HMI tags "Default tag table"
   "Tag_ScreenNumber" : UInt AT %DB1.DBW0
   "Part At Entry (NC)" : Bool AT %DB1.DBX0.0
   "InputsDB_Sensors_Part Entry" : Bool = PLC InputsDB.Sensors."Part Entry" AT %DB1.DBX0.0, 100 ms
   "Modes_Modes_RunMode" : Bool = PLC Modes.Modes.RunMode, 100 ms
   "HmiDb_ActivateUnloadHmi" : Bool = PLC HmiDb.HmiModes.ActivateUnloadHmi, 100 ms
   "Modes_Modes_StopMode" : Bool = PLC Modes.Modes.StoppestMode, 100 ms
   "Modes_Modes_ResetMode" : Bool = PLC Modes.Modes.ResetMode, 100 ms
   "HmiDb_HmiRunMode" : Bool = PLC HmiDb.HmiModes.HmiRunMode, 100 ms
   "HmiDb_HmiStopmode" : Bool = PLC HmiDb.HmiModes.HmiStopmode, 100 ms
   "HmiDb_HmiResetMode" : Bool = PLC HmiDb.HmiModes.HmiResetMode, 100 ms
   "InputsDB_Sensors_Part Load" : Bool = PLC InputsDB.Sensors."Part Load", 100 ms
   "InputsDB_Sensors_Part Unload" : Bool = PLC InputsDB.Sensors."Part Unload", 100 ms
   "InputsDB_Sensors_Part Exit" : Bool = PLC InputsDB.Sensors."Part Exit", 100 ms
   "InputsDB_Sensors_Crane Default" : Bool = PLC InputsDB.Sensors."Crane Default", 100 ms
   "InputsDB_Sensors_Crane Entry" : Bool = PLC InputsDB.Sensors."Crane Entry", 100 ms
   "InputsDB_Sensors_Color Sensor" : Int = PLC InputsDB.Sensors."Color Sensor", 100 ms
   "Modes_SafetyStops_ProductionStop" : Bool = PLC Modes.StopMethods.ProductionStop, 100 ms
   "Modes_SafetyStops_SafetyStop" : Bool = PLC Modes.StopMethods.SafetyStop, 100 ms
   "alarmStuck" : Int = PLC alarmStuck AT %QW34, 100 ms
   "alarmreceivedstuck" : UInt, internal
   "alarmLoaderFull" : Int = PLC alarmLoaderFull AT %QW36, 100 ms
   "alarmUnloaderEmpty" : Int = PLC alarmUnloaderEmpty AT %QW38, 100 ms
   "Modes_JogMode" : Bool = PLC Modes.Modes.JogMode, 100 ms
   "HmiDb_HmiRunEntryConv" : Bool = PLC HmiDb.ActivateAcutator.HmiRunEntryConv, 100 ms
   "HmiDb_HmiRunExitConv" : Bool = PLC HmiDb.ActivateAcutator.HmiRunExitConv, 100 ms
   "EntryConv" : Int = PLC InputsDB.ConvertedConveyors.EntryConvSensorVal, 100 ms
   "LoadingConv" : Int = PLC InputsDB.ConvertedConveyors.LoadingConvSensorVal, 100 ms
   "UnloadingConv" : Int = PLC InputsDB.ConvertedConveyors.UnloadingSensorVal, 100 ms
   "ExitConv" : Int = PLC InputsDB.ConvertedConveyors.ExitConvSensorVal, 100 ms
   "ohioselecter" : Int AT %DB1.DBW0
   "unloadingms" : Real = PLC InputsDB.ConvertedConveyors.UnloadingScaleX, 100 ms
   "loadingms" : Real = PLC InputsDB.ConvertedConveyors.LoadingConvScalex, 100 ms
   "exitms" : Real = PLC InputsDB.ConvertedConveyors.ExitConvScaleX, 100 ms
   "entryms" : Real = PLC InputsDB.ConvertedConveyors.EntryConvScalex, 100 ms
   "OutputsDB_CraneOutput_XScalex" : Int = PLC OutputsDB.CraneOutput.Xmm, 100 ms
   "OutputsDB_CraneOutput_YScalex" : Int = PLC OutputsDB.CraneOutput.Ymm, 100 ms
   "HmiDb_HmiExtendExit" : Bool = PLC HmiDb.ActivateAcutator.HmiExtendExit, 100 ms
   "HmiDb_HmiExtendEntry" : Bool = PLC HmiDb.ActivateAcutator.HmiExtendEntry, 100 ms
   "InputsDB_Sensors_Crane Exit" : Bool = PLC InputsDB.Sensors."Crane Exit", 100 ms
   "InputsDB_ConveyorCalibrationBarSlider" : Int = PLC InputsDB.ConveyorCalibrationBarSlider, 100 ms
   "InputsDB_ConveyorCalibrationPicker" : Int = PLC InputsDB.ConveyorCalibrationPicker, 100 ms
   "InputsDB_ConveyorSaveCalVal_HmiDisplayMin" : Int = PLC InputsDB.ConveyorSaveCalVal.Min.HmiDisplayMin, 100 ms
   "InputsDB_ConveyorSaveCalVal_HmiDisplayMax" : Int = PLC InputsDB.ConveyorSaveCalVal.Max.HmiDisplayMax, 100 ms
   "InputsDB_ConveyorSaveCalVal_ActualdisplayMax" : Int = PLC InputsDB.ConveyorSaveCalVal.Max.ActualdisplayMax, 100 ms
   "InputsDB_ConveyorSaveCalVal_ActualdisplayMin" : Int = PLC InputsDB.ConveyorSaveCalVal.Min.ActualdisplayMin, 100 ms
   "InputsDB_ConveyorSaveCalVal_Save" : Bool = PLC InputsDB.ConveyorSaveCalVal.Save, 100 ms
   "InputsDB_ConveyorSaveCalVal_DisplayMm/s" : Real = PLC InputsDB.ConveyorSaveCalVal.DisplayMm/s, 100 ms
   "jogmodeDB_CraneXjog" : Int = PLC jogmodeDB.CraneXjog, 100 ms
   "jogmodeDB_CraneYjog" : Int = PLC jogmodeDB.CraneYjog, 100 ms
   "HmiDb_Static_1_HmiOrderAmount" : Int = PLC HmiDb.HmiOrderMode.HmiOrderAmount, 100 ms
   "HmiDb_Static_1_HmiColorSelected" : Int = PLC HmiDb.HmiOrderMode.HmiColorSelected, 100 ms
   "HmiDb_Static_1_HmiExecuteOrder" : Bool = PLC HmiDb.HmiOrderMode.HmiExecuteOrder, 100 ms
   "Crane Current Z Position" : Int = PLC "Crane Current Z Position" AT %IW28, 100 ms
   "HmiDb_ActivateAcutator_hmilighttest" : Bool = PLC HmiDb.ActivateAcutator.hmilighttest, 100 ms
   "activateloadconv" : Bool = PLC HmiDb.ActivateAcutator.HmiRunLoadConv, 100 ms
   "activateunloadconv" : Bool = PLC HmiDb.ActivateAcutator.HmiRunUnloadConv, 100 ms
   "Reset Button" : Bool = PLC "Reset Button" AT %I0.1, 100 ms
   "Start Button" : Bool = PLC "Start Button" AT %I0.0, 100 ms
   "Stop Button (NC)" : Bool = PLC "Stop Button (NC)" AT %I0.2, 100 ms
   "adminornot" : Bool AT %DB1.DBX0.0
   "userid" : Int, internal
   "Modes_Sequences_SequenceLoader" : Int = PLC Modes.Sequences.SequenceLoader, 100 ms

discrete alarms
   1: 'Verkar att ha fastnat', class Errors, trigger "alarmreceivedstuck" bit 0
   2: 'Kan inte lasta fler pga. fullt', class Warnings, trigger "alarmLoaderFull" bit 0
   3: 'Kan inte last ur pga. tomt', class Warnings, trigger "alarmUnloaderEmpty" bit 0

analog alarms
   1: '', class Errors, trigger "Crane Current Z Position"

text list "conveyorpicker": 0..1 'entry'; 2..3 'exit'; 4..5 'load'; 6..7 'unload'

text list "ColorBoxList": 0..1 'Gray'; 2..3 'Blue'; 4..5 'Green'

screen "Main" 800x480
   Button "Button_1" at 22,109 size 123x50; TextOff 'Run Mode'
      Appearance <- "Modes_Modes_RunMode"
      on Press: SetBit("HmiDb_HmiRunMode")
      on Release: ResetBit("HmiDb_HmiRunMode")
   Button "Button_2" at 22,221 size 123x50; TextOff 'Reset Mode'
      Appearance <- "Modes_Modes_ResetMode"
      on Press: SetBit("HmiDb_HmiResetMode")
      on Release: ResetBit("HmiDb_HmiResetMode")
   Button "Button_3" at 22,164 size 123x50; TextOff 'Stop Mode'
      on Press: SetBit("HmiDb_HmiStopmode")
      on Release: ResetBit("HmiDb_HmiStopmode")
      Appearance <- "Modes_Modes_StopMode"
   Button "Button_4" at 280,336 size 149x50; TextOff 'Safety Stop'
      on Click: InvertBit("Modes_SafetyStops_SafetyStop"); InvertBit("Modes_SafetyStops_ProductionStop")
      Appearance <- "Modes_SafetyStops_SafetyStop"
   Button "Button_5" at 499,336 size 149x50; TextOff 'Production Stop'
      on Click: InvertBit("Modes_SafetyStops_ProductionStop"); InvertBit("Modes_SafetyStops_SafetyStop")
      Appearance <- "Modes_SafetyStops_ProductionStop"
   Button "Button_6" at 22,336 size 123x50; TextOff 'Unload Mode'
      Appearance <- "HmiDb_ActivateUnloadHmi"
      on Click: InvertBit("HmiDb_ActivateUnloadHmi")
   SymbolicIOField "Symbolic I/O field_1" at 595,8 size 170x32; TextOff '0'; TextOn '1'; TextList "TextList_ScreenNames"
      ProcessValue <- "ohioselecter"
      on Change: ActivateScreenByNumber("ohioselecter", 0)
      Visibility <- "userid"
   Button "Button_7" at 22,8 size 96x32; TextOff 'Log Out'
      on Activate: function_f23ef4c9()
      on Change: ActivateScreen("Login", 0)

screen "JogMode" 800x480, template "Template_1"
   on GenerateScreen: SetTag("Tag_ScreenNumber", 1)
   Button "Button_1" at 17,61 size 168x32; TextOff 'Test Lights'
      on Click: InvertBit("HmiDb_ActivateAcutator_hmilighttest")
      Appearance <- "HmiDb_ActivateAcutator_hmilighttest"
   Button "Button_2" at 17,109 size 167x32; TextOff 'Extend Crane Entry'
      on Click: InvertBit("HmiDb_HmiExtendEntry")
      Appearance <- "HmiDb_HmiExtendEntry"
   Button "Button_3" at 17,155 size 167x32; TextOff 'Extend Crane Exit'
      on Click: InvertBit("HmiDb_HmiExtendExit")
      Appearance <- "HmiDb_HmiExtendExit"
   Button "Button_4" at 18,204 size 167x32; TextOff 'Entry Conveyor'
      on Click: InvertBit("HmiDb_HmiRunEntryConv")
      Appearance <- "HmiDb_HmiRunEntryConv"
   Button "Button_5" at 18,256 size 167x32; TextOff 'Exit Conveyor'
      on Click: InvertBit("HmiDb_HmiRunExitConv")
      Appearance <- "HmiDb_HmiRunExitConv"
   Button "Button_8" at 18,306 size 167x32; TextOff 'Load Conveyor'
      on Click: InvertBit("activateloadconv")
      Appearance <- "activateloadconv"
   Button "Button_9" at 262,428 size 260x32; TextOff 'Jog Mode'
      on Click: InvertBit("Modes_JogMode")
      Appearance <- "Modes_JogMode"
      on Deactivate: ResetBit("HmiDb_ActivateAcutator_hmilighttest"); ResetBit("HmiDb_HmiExtendEntry"); ResetBit("HmiDb_HmiExtendExit"); ResetBit("HmiDb_HmiRunExitConv"); ResetBit("HmiDb_HmiRunEntryConv"); ResetBit("activateloadconv"); ResetBit("activateunloadconv"); SetTag("jogmodeDB_CraneXjog", 0); SetTag("jogmodeDB_CraneYjog", 0)
      on Activate: ResetBit("HmiDb_ActivateAcutator_hmilighttest"); ResetBit("HmiDb_HmiExtendEntry"); ResetBit("HmiDb_HmiExtendExit"); ResetBit("HmiDb_HmiRunExitConv"); ResetBit("HmiDb_HmiRunEntryConv"); ResetBit("activateloadconv"); ResetBit("activateunloadconv"); SetTag("jogmodeDB_CraneXjog", 0); SetTag("jogmodeDB_CraneYjog", 0)
   Group "Group" at 594,43 size 185x38
   Group "Group_1" at 594,82 size 185x38
   Group "Group_2" at 594,121 size 185x38
   Group "Group_3" at 594,161 size 185x38
   Group "Group_4" at 594,201 size 185x38
   Group "Group_5" at 594,319 size 185x38
   Group "Group_6" at 594,240 size 185x38
   Group "Group_7" at 594,279 size 185x38
   SymbolicIOField "Symbolic I/O field_1" at 595,8 size 170x32; TextOn '1'; TextOff '0'; TextList "TextList_ScreenNames"
      on Change: ActivateScreenByNumber("ohioselecter", 0)
      ProcessValue <- "ohioselecter"
   Slider "Slider_2" at 262,61 size 80x329; Caption 'SIMATIC'
      ProcessValue <- "jogmodeDB_CraneXjog"
   Slider "Slider_1" at 439,61 size 80x328; Caption 'SIMATIC'
      ProcessValue <- "jogmodeDB_CraneYjog"
   Button "Button_6" at 18,355 size 167x32; TextOff 'Unload Conveyor'
      on Click: InvertBit("activateunloadconv")
      Appearance <- "activateunloadconv"
   Group "Group_8" at 595,359 size 185x38
   Group "Group_9" at 594,399 size 185x38
   Group "Group_10" at 595,439 size 185x38
   TextField "Text field_12" at 288,20 size 17x23; Text 'X'
   TextField "Text field_13" at 468,20 size 17x23; Text 'Y'
   Circle "Circle_3" at 741,43 size 37x37
      Appearance <- "InputsDB_Sensors_Part Entry"
   TextField "Text field_1" at 618,53 size 110x23; Text 'Part at Entry'
   Circle "Circle_6" at 741,82 size 37x37
      Appearance <- "InputsDB_Sensors_Part Load"
   TextField "Text field_2" at 618,92 size 108x23; Text 'Part At Load'
   Circle "Circle_9" at 741,121 size 37x37
      Appearance <- "InputsDB_Sensors_Part Unload"
   TextField "Text field_3" at 618,131 size 126x23; Text 'Part At Unload'
   Circle "Circle_12" at 741,161 size 37x37
      Appearance <- "InputsDB_Sensors_Part Exit"
   TextField "Text field_4" at 618,171 size 101x23; Text 'Part At Exit'
   Circle "Circle_15" at 741,201 size 37x37
      Appearance <- "InputsDB_Sensors_Crane Default"
   TextField "Text field_5" at 618,211 size 118x23; Text 'Crane Default'
   Circle "Circle_18" at 741,319 size 37x37
      Appearance <- "InputsDB_Sensors_Color Sensor"
   TextField "Text field_6" at 618,329 size 120x23; Text 'Color Sensor'
   Circle "Circle_21" at 741,240 size 37x37
      Appearance <- "InputsDB_Sensors_Crane Exit"
   TextField "Text field_7" at 618,250 size 114x23; Text 'Crane At Exit'
   Circle "Circle_24" at 741,279 size 37x37
      Appearance <- "InputsDB_Sensors_Crane Entry"
   TextField "Text field_8" at 618,289 size 125x23; Text 'Crane At Entry'
   Circle "Circle_27" at 742,359 size 37x37
      Appearance <- "Start Button"
   TextField "Text field_9" at 619,369 size 132x23; Text 'Green Button'
   Circle "Circle_30" at 741,399 size 37x37
      Appearance <- "Stop Button (NC)"
   TextField "Text field_10" at 618,409 size 113x23; Text 'Red Button'
   Circle "Circle_33" at 742,439 size 37x37
      Appearance <- "Reset Button"
   TextField "Text field_11" at 619,449 size 118x23; Text 'Blue Button'

screen "larm" 800x480, template "Template_1"
   on GenerateScreen: SetTag("Tag_ScreenNumber", 0)
   AlarmView "Alarm view_1" at 0,52 size 799x427
   SymbolicIOField "Symbolic I/O field_1" at 595,8 size 170x32; TextOn '1'; TextOff '0'; TextList "TextList_ScreenNames"
      on Change: ActivateScreenByNumber("ohioselecter", 4)
      ProcessValue <- "ohioselecter"

screen "CalibrationConveyor" 800x480
   on GenerateScreen: SetTag("Tag_ScreenNumber", 2)
   Slider "Slider_4" at 402,135 size 80x230; Caption 'SIMATIC'
      ProcessValue <- "InputsDB_ConveyorCalibrationBarSlider"
   SymbolicIOField "Symbolic I/O field_1" at 595,8 size 170x32; TextOn '1'; TextOff '0'; TextList "TextList_ScreenNames"
      on Change: ActivateScreenByNumber("ohioselecter", 0)
      ProcessValue <- "ohioselecter"
   Bar "Bar_2" at 341,135 size 61x230; MinimumValue 0; MaximumValue 100
      MaximumValue <- "InputsDB_ConveyorSaveCalVal_ActualdisplayMax"
      MinimumValue <- "InputsDB_ConveyorSaveCalVal_ActualdisplayMin"
      ProcessValue <- "InputsDB_ConveyorSaveCalVal_DisplayMm/s"
   SymbolicIOField "Symbolic I/O field_2" at 595,75 size 170x32; TextOff '0'; TextOn '1'; TextList "conveyorpicker"
      ProcessValue <- "InputsDB_ConveyorCalibrationPicker"
   IOField "I/O field_1" at 274,75 size 100x32; FormatPattern 99999
      ProcessValue <- "InputsDB_ConveyorSaveCalVal_HmiDisplayMin"
   IOField "I/O field_2" at 440,75 size 99x32; FormatPattern 99999
      ProcessValue <- "InputsDB_ConveyorSaveCalVal_HmiDisplayMax"
   TextField "Text field_1" at 306,40 size 37x23; Text 'Min'
   TextField "Text field_2" at 469,37 size 42x23; Text 'Max'
   Button "Button_1" at 305,380 size 225x49; TextOff 'Save'
      on Press: InvertBit("InputsDB_ConveyorSaveCalVal_Save")
      on Release: InvertBit("InputsDB_ConveyorSaveCalVal_Save")

screen "Login" 800x480
   Button "Button_1" at 316,188 size 198x108; TextOff 'Login'
      on Activate: function_a2a04561()
      on Change: ActivateScreen("Main", 0)

scheduled task "Task_1"
   on Action: function_e1ab61de("userid")
*)

(* ===== HMI "HMI_RT_2" =====
system functions are stored by id; their names below are inferred from use
connection "HMI_Connection_2": ETHERNET, S7_1500_OMS
connection "HMI_Connection_3": ETHERNET, S7_1500_OMS

HMI tags "Default tag table"
   "HmiDb_Static_1_HmiOrderAmount" : Int = PLC HmiDb.HmiOrderMode.HmiOrderAmount, 1 s
   "HmiDb_Static_1_HmiColorSelected" : Int = PLC HmiDb.HmiOrderMode.HmiColorSelected, 1 s
   "ohioselecter" : Int AT %DB1.DBW0
   "HmiDb_Static_1_HmiExecuteOrder" : Bool = PLC HmiDb.HmiOrderMode.HmiExecuteOrder, 1 s
   "InputsDB_ErrorStuck" : Bool = PLC InputsDB.ErrorStuck, 1 s
   "pause" : Bool = PLC HmiDb.HmiOrderMode.HmiPauseOrder, 1 s
   "THEscreen" : Int AT %DB1.DBW0
   "Modes_Modes_RunMode" : Bool = PLC Modes.Modes.RunMode, 1 s
   "Modes_Modes_StoppestMode" : Bool = PLC Modes.Modes.StoppestMode, 1 s
   "Modes_Modes_ResetMode" : Bool = PLC Modes.Modes.ResetMode, 1 s
   "Modes_Modes_Unloadmode" : Bool = PLC Modes.Modes.Unloadmode, 1 s
   "ColorCounterDB_Gray" : Int = PLC ColorDB.Gray, 1 s
   "ColorCounterDB_Blue" : Int = PLC ColorDB.Blue, 100 ms
   "ColorCounterDB_Green" : Int = PLC ColorDB.Green, 1 s
   "InputsDB_RunArmX" : Bool = PLC InputsDB.Crane.RunArmX, 1 s
   "InputsDB_RunArmY" : Bool = PLC InputsDB.Crane.RunArmY, 1 s
   "InputsDB_RunEntryConveyor" : Bool = PLC InputsDB.RunConveyor.RunEntryConveyor, 1 s
   "InputsDB_RunLoadingConveyor" : Bool = PLC InputsDB.RunConveyor.RunLoadingConveyor, 1 s
   "InputsDB_RunUnloadingConveyor" : Bool = PLC InputsDB.RunConveyor.RunUnloadingConveyor, 1 s
   "InputsDB_RunExitConveyor" : Bool = PLC InputsDB.RunConveyor.RunExitConveyor, 1 s
   "InputsDB_YisMoving" : Bool = PLC InputsDB.YisMoving, 1 s
   "InputsDB_XisMoving" : Bool = PLC InputsDB.XisMoving, 1 s
   "OutputsDB_MoveForkEntryLoad" : Bool = PLC OutputsDB.ForkController.MoveForkEntryLoad, 1 s
   "OutputsDB_MoveForkExitLoad" : Bool = PLC OutputsDB.ForkController.MoveForkExitLoad, 1 s
   "coolboxmover" : Int = PLC HmiDb.BoxyMover, 1 s
   "coolboxmover2" : Int = PLC HmiDb.BoxyMover2 AT %DB1.DBW0, 1 s
   "HmiDb_BoxyMover2" : Int = PLC HmiDb.BoxyMover2, 1 s
   "HmiDb_ClearStock" : Bool = PLC HmiDb.ClearStock, 1 s
   "HmiDb_ClearCounter" : Bool = PLC HmiDb.ClearCounter, 1 s
   "xlist" : Int = PLC HmiDb.XListColumn, 1 s
   "ylist" : Int = PLC HmiDb.YListColumn, 1 s
   "HmiDb_HmiSaveArmCal" : Bool = PLC HmiDb.HmiSaveArmCalX, 1 s
   "HmiDb_HmiSaveArmCalY" : Bool = PLC HmiDb.HmiSaveArmCalY, 1 s
   "HmiDb_CalInputVal" : Int = PLC HmiDb.CalInputVal, 100 ms
   "HmiDb_CurrentPositionX" : Int = PLC HmiDb.CurrentPositionX, 100 ms
   "HmiDb_CurrentPositionY" : Int = PLC HmiDb.CurrentPositionY, 100 ms
   "HmiDb_oke" : String[254] = PLC HmiDb.oke, 1 s
   "InputsDB_FreeSlotCounter" : Int = PLC InputsDB.FreeSlotCounter, 1 s
   "IEC_Counter_0_DB_5_PV" : Int = PLC FreeSlotCounter.PV, 1 s
   "InputsDB_totalcounter" : Int = PLC InputsDB.totalcounter, 1 s
   "InputsDB_totalremovedcounter" : Int = PLC InputsDB.totalremovedcounter, 1 s
   "AlreadyFilledSlotArray_Row1Y{0}" : Int = PLC AlreadyFilledSlotArray.Row1Y[0], 1 s
   "AlreadyFilledSlotArray_Row2Y{0}" : Int = PLC AlreadyFilledSlotArray.Row2Y[0], 1 s
   "AlreadyFilledSlotArray_Row3Y{0}" : Int = PLC AlreadyFilledSlotArray.Row3Y[0], 1 s
   "AlreadyFilledSlotArray_Row4Y{0}" : Int = PLC AlreadyFilledSlotArray.Row4Y[0], 1 s
   "AlreadyFilledSlotArray_Row5Y{0}" : Int = PLC AlreadyFilledSlotArray.Row5Y[0], 1 s
   "AlreadyFilledSlotArray_Row6Y{0}" : Int = PLC AlreadyFilledSlotArray.Row6Y[0], 1 s
   "AlreadyFilledSlotArray_Row7Y{0}" : Int = PLC AlreadyFilledSlotArray.Row7Y[0], 1 s
   "AlreadyFilledSlotArray_Row8Y{0}" : Int = PLC AlreadyFilledSlotArray.Row8Y[0], 1 s
   "AlreadyFilledSlotArray_Row9Y{0}" : Int = PLC AlreadyFilledSlotArray.Row9Y[0], 1 s
   "AlreadyFilledSlotArray_Row1Y{1}" : Int = PLC AlreadyFilledSlotArray.Row1Y[1], 1 s
   "AlreadyFilledSlotArray_Row2Y{1}" : Int = PLC AlreadyFilledSlotArray.Row2Y[1], 1 s
   "AlreadyFilledSlotArray_Row3Y{1}" : Int = PLC AlreadyFilledSlotArray.Row3Y[1], 1 s
   "AlreadyFilledSlotArray_Row4Y{1}" : Int = PLC AlreadyFilledSlotArray.Row4Y[1], 1 s
   "AlreadyFilledSlotArray_Row5Y{1}" : Int = PLC AlreadyFilledSlotArray.Row5Y[1], 1 s
   "AlreadyFilledSlotArray_Row6Y{1}" : Int = PLC AlreadyFilledSlotArray.Row6Y[1], 1 s
   "AlreadyFilledSlotArray_Row7Y{1}" : Int = PLC AlreadyFilledSlotArray.Row7Y[1], 1 s
   "AlreadyFilledSlotArray_Row8Y{1}" : Int = PLC AlreadyFilledSlotArray.Row8Y[1], 1 s
   "AlreadyFilledSlotArray_Row9Y{1}" : Int = PLC AlreadyFilledSlotArray.Row9Y[1], 1 s
   "AlreadyFilledSlotArray_Row9Y{2}" : Int = PLC AlreadyFilledSlotArray.Row9Y[2], 1 s
   "AlreadyFilledSlotArray_Row8Y{2}" : Int = PLC AlreadyFilledSlotArray.Row8Y[2], 1 s
   "AlreadyFilledSlotArray_Row7Y{2}" : Int = PLC AlreadyFilledSlotArray.Row7Y[2], 1 s
   "AlreadyFilledSlotArray_Row6Y{2}" : Int = PLC AlreadyFilledSlotArray.Row6Y[2], 1 s
   "AlreadyFilledSlotArray_Row5Y{2}" : Int = PLC AlreadyFilledSlotArray.Row5Y[2], 1 s
   "AlreadyFilledSlotArray_Row4Y{2}" : Int = PLC AlreadyFilledSlotArray.Row4Y[2], 1 s
   "AlreadyFilledSlotArray_Row3Y{2}" : Int = PLC AlreadyFilledSlotArray.Row3Y[2], 1 s
   "AlreadyFilledSlotArray_Row2Y{2}" : Int = PLC AlreadyFilledSlotArray.Row2Y[2], 1 s
   "AlreadyFilledSlotArray_Row1Y{2}" : Int = PLC AlreadyFilledSlotArray.Row1Y[2], 1 s
   "AlreadyFilledSlotArray_Row9Y{3}" : Int = PLC AlreadyFilledSlotArray.Row9Y[3], 1 s
   "AlreadyFilledSlotArray_Row8Y{3}" : Int = PLC AlreadyFilledSlotArray.Row8Y[3], 1 s
   "AlreadyFilledSlotArray_Row7Y{3}" : Int = PLC AlreadyFilledSlotArray.Row7Y[3], 1 s
   "AlreadyFilledSlotArray_Row6Y{3}" : Int = PLC AlreadyFilledSlotArray.Row6Y[3], 1 s
   "AlreadyFilledSlotArray_Row5Y{3}" : Int = PLC AlreadyFilledSlotArray.Row5Y[3], 1 s
   "AlreadyFilledSlotArray_Row4Y{3}" : Int = PLC AlreadyFilledSlotArray.Row4Y[3], 1 s
   "AlreadyFilledSlotArray_Row3Y{3}" : Int = PLC AlreadyFilledSlotArray.Row3Y[3], 1 s
   "AlreadyFilledSlotArray_Row2Y{3}" : Int = PLC AlreadyFilledSlotArray.Row2Y[3], 1 s
   "AlreadyFilledSlotArray_Row1Y{3}" : Int = PLC AlreadyFilledSlotArray.Row1Y[3], 1 s
   "AlreadyFilledSlotArray_Row1Y{4}" : Int = PLC AlreadyFilledSlotArray.Row1Y[4], 1 s
   "AlreadyFilledSlotArray_Row2Y{4}" : Int = PLC AlreadyFilledSlotArray.Row2Y[4], 1 s
   "AlreadyFilledSlotArray_Row3Y{4}" : Int = PLC AlreadyFilledSlotArray.Row3Y[4], 1 s
   "AlreadyFilledSlotArray_Row4Y{4}" : Int = PLC AlreadyFilledSlotArray.Row4Y[4], 1 s
   "AlreadyFilledSlotArray_Row5Y{4}" : Int = PLC AlreadyFilledSlotArray.Row5Y[4], 1 s
   "AlreadyFilledSlotArray_Row6Y{4}" : Int = PLC AlreadyFilledSlotArray.Row6Y[4], 1 s
   "AlreadyFilledSlotArray_Row7Y{4}" : Int = PLC AlreadyFilledSlotArray.Row7Y[4], 1 s
   "AlreadyFilledSlotArray_Row8Y{4}" : Int = PLC AlreadyFilledSlotArray.Row8Y[4], 1 s
   "AlreadyFilledSlotArray_Row9Y{4}" : Int = PLC AlreadyFilledSlotArray.Row9Y[4], 1 s
   "AlreadyFilledSlotArray_Row9Y{5}" : Int = PLC AlreadyFilledSlotArray.Row9Y[5], 1 s
   "AlreadyFilledSlotArray_Row8Y{5}" : Int = PLC AlreadyFilledSlotArray.Row8Y[5], 1 s
   "AlreadyFilledSlotArray_Row7Y{5}" : Int = PLC AlreadyFilledSlotArray.Row7Y[5], 1 s
   "AlreadyFilledSlotArray_Row6Y{5}" : Int = PLC AlreadyFilledSlotArray.Row6Y[5], 1 s
   "AlreadyFilledSlotArray_Row5Y{5}" : Int = PLC AlreadyFilledSlotArray.Row5Y[5], 1 s
   "AlreadyFilledSlotArray_Row4Y{5}" : Int = PLC AlreadyFilledSlotArray.Row4Y[5], 1 s
   "AlreadyFilledSlotArray_Row3Y{5}" : Int = PLC AlreadyFilledSlotArray.Row3Y[5], 1 s
   "AlreadyFilledSlotArray_Row2Y{5}" : Int = PLC AlreadyFilledSlotArray.Row2Y[5], 1 s
   "AlreadyFilledSlotArray_Row1Y{5}" : Int = PLC AlreadyFilledSlotArray.Row1Y[5], 1 s
   "OutputsDB_CraneOutput_Xmm" : Int = PLC OutputsDB.CraneOutput.Xmm, 1 s
   "OutputsDB_CraneOutput_Ymm" : Int = PLC OutputsDB.CraneOutput.Ymm, 1 s
   "Modes_Modes_JogMode" : Bool = PLC Modes.Modes.JogMode, 1 s
   "jogmodeDB_CraneXjog" : Int = PLC jogmodeDB.CraneXjog, 1 s
   "jogmodeDB_CraneYjog" : Int = PLC jogmodeDB.CraneYjog, 1 s
   "InputsDB_AdjustX" : Int = PLC InputsDB.AdjustX, 1 s
   "InputsDB_PressAdjustX" : Bool = PLC InputsDB.PressAdjustX, 1 s
   "InputsDB_AdjustY" : Int = PLC InputsDB.AdjustY, 1 s
   "InputsDB_PressAdjustY" : Bool = PLC InputsDB.PressAdjustY, 1 s
   "HmiDb_HmiOrderMode_OrderDelivered" : Int = PLC HmiDb.HmiOrderMode.OrderDelivered, 1 s

text list "scadascreenlist": 1 'Order Screen'; 2 'Status Screen'; 3 'Calibrate Screen'

text list "ColorBoxList": 0..1 'Gray'; 2..3 'Blue'; 4..5 'Green'

text list "coolgraphics": 0..1 ''

text list "XarrayList": 0 'Column 1 X'; 1 'Column 2 X'; 2 'Column 3 X'; 3 'Column 4 X'; 4 'Column 5 X'; 5 'Column 6 X'; 6 'Column 7 X'; 7 'Column 8 X'; 8 'Column 9 X'

text list "ZarrayList": 0 'Column 1 Z'; 1 'Column 2 Z'; 2 'Column 3 Z'; 3 'Column 4 Z'; 4 'Column 5 Z'; 5 'Column 6 Z'

graphic list "XaxisMotor": 0..1 'Graphic_2'; 2..3 'Graphic_3'; 4..5 'Graphic_4'; 6..7 'Graphic_5'

graphic list "ZaxisMotor": 0..1 'Graphic_2'; 2..3 'Graphic_3'; 4..5 'Graphic_4'; 6..7 'Graphic_5'

screen "Order" 800x600
   TextField "Text field_1" at 306,56 size 170x34; Text 'Order Screen'
   IOField "I/O field_1" at 67,178 size 122x32; FormatPattern 9999
      ProcessValue <- "HmiDb_Static_1_HmiOrderAmount"
   TextField "Text field_2" at 68,147 size 120x23; Text 'Order Amount'
   Button "Button_1" at 465,192 size 96x32; TextOff 'Execute'
      on Release: InvertBit("HmiDb_Static_1_HmiExecuteOrder")
      on Press: InvertBit("HmiDb_Static_1_HmiExecuteOrder")
   TextField "Text field_3" at 250,147 size 99x23; Text 'Order Color'
   SymbolicIOField "Symbolic I/O field_2" at 218,178 size 170x32; TextOn '1'; TextOff '0'; TextList "ColorBoxList"
      ProcessValue <- "HmiDb_Static_1_HmiColorSelected"
   Button "Button_2" at 578,192 size 96x32; TextOff 'Pause'
      on Press: InvertBit("pause")
      on Release: InvertBit("pause")
   SymbolicIOField "Symbolic I/O field_1" at 595,8 size 170x32; TextOn '1'; TextOff '0'; TextList "scadascreenlist"
      on Change: ActivateScreenByNumber("THEscreen", 0)
      ProcessValue <- "THEscreen"
   IOField "I/O field_2" at 66,246 size 122x32; FormatPattern 9999
      ProcessValue <- "HmiDb_HmiOrderMode_OrderDelivered"
   TextField "Text field_4" at 63,217 size 152x23; Text 'Delivered Amount'

screen "Status" 800x600
   SymbolicIOField "Symbolic I/O field_1" at 595,8 size 170x32; TextOn '1'; TextOff '0'; TextList "scadascreenlist"
      on Change: ActivateScreenByNumber("THEscreen", 1)
      ProcessValue <- "THEscreen"
   TextField "Text field_1" at 646,187 size 129x39; Text 'Running'
   TextField "Text field_2" at 646,251 size 124x39; Text 'Stopped'
   TextField "Text field_3" at 644,187 size 129x39; Text 'Running'
      Appearance <- "Modes_Modes_RunMode"
   TextField "Text field_4" at 644,251 size 124x39; Text 'Stopped'
      Appearance <- "Modes_Modes_StoppestMode"
   TextField "Text field_5" at 646,307 size 145x39; Text 'Resetting'
   TextField "Text field_6" at 644,307 size 145x39; Text 'Resetting'
      Appearance <- "Modes_Modes_ResetMode"
   TextField "Text field_7" at 512,372 size 153x39; Text 'Unloading'
   TextField "Text field_8" at 510,372 size 153x39; Text 'Unloading'
      Appearance <- "Modes_Modes_Unloadmode"
   TextField "Text field_9" at 673,373 size 121x39; Text 'Loading'
   TextField "Text field_10" at 671,373 size 121x39; Text 'Loading'
      Appearance <- "Modes_Modes_Unloadmode"
   TextField "Text field_11" at 554,454 size 90x22; Text 'Gray Boxes'
   TextField "Text field_12" at 555,498 size 87x22; Text 'Blue Boxes'
   TextField "Text field_13" at 549,538 size 99x22; Text 'Green Boxes'
   IOField "I/O field_1" at 679,454 size 96x31; FormatPattern 9999
      ProcessValue <- "ColorCounterDB_Gray"
   IOField "I/O field_2" at 679,497 size 96x31; FormatPattern 9999
      ProcessValue <- "ColorCounterDB_Blue"
   IOField "I/O field_3" at 678,538 size 96x31; FormatPattern 9999
      ProcessValue <- "ColorCounterDB_Green"
   SymbolLibrary "Symbol library_8" at 530,84 size 94x89
   SymbolLibrary "Symbol library_5" at 40,477 size 120x109
      Appearance <- "InputsDB_RunEntryConveyor"
   SymbolLibrary "Symbol library_6" at 40,370 size 120x109
      Appearance <- "InputsDB_RunLoadingConveyor"
   SymbolLibrary "Symbol library_3" at 40,132 size 120x120
      Appearance <- "InputsDB_RunUnloadingConveyor"
   SymbolLibrary "Symbol library_4" at 40,12 size 120x120
      Appearance <- "InputsDB_RunExitConveyor"
   SymbolLibrary "Symbol library_7" at 530,86 size 94x89
      Visibility <- "OutputsDB_MoveForkEntryLoad"
   SymbolLibrary "Symbol library_9" at 530,85 size 94x89
      Visibility <- "OutputsDB_MoveForkExitLoad"
   SymbolLibrary "Symbol library_1" at 262,369 size 34x97
      Appearance <- "InputsDB_YisMoving"
   SymbolLibrary "Symbol library_2" at 214,520 size 97x34
      Appearance <- "InputsDB_XisMoving"
   GraphicView "Graphic view_1" at 352,491 size 149x97; Picture "Graphic_2"
      Visibility <- "InputsDB_RunArmX"
   GraphicView "Graphic view_2" at 352,491 size 149x97; Picture "Graphic_3"
      Visibility <- "InputsDB_RunArmX"
   GraphicView "Graphic view_4" at 352,376 size 149x97; Picture "Graphic_2"
      Visibility <- "InputsDB_RunArmY"
   GraphicView "Graphic view_5" at 352,376 size 149x97; Picture "Graphic_3"
      Visibility <- "InputsDB_RunArmY"
   SymbolLibrary "Symbol library_10" at 251,520 size 97x34
      Appearance <- "InputsDB_XisMoving"
   SymbolLibrary "Symbol library_11" at 263,406 size 34x97
      Appearance <- "InputsDB_YisMoving"
   SymbolLibrary "Symbol library_13" at 58,493 size 83x83
      VerticalMovement <- "coolboxmover"
      Visibility <- "coolboxmover"
   SymbolLibrary "Symbol library_12" at 56,159 size 83x83
      VerticalMovement <- "coolboxmover2"
      Visibility <- "HmiDb_BoxyMover2"
   Button "Button_1" at 516,219 size 119x32; TextOff 'Clear Stock'
      on Press: function_efd93a16("Pop-up screen_1", 0, 0, -1, -1, 1)
   Button "Button_2" at 516,290 size 119x32; TextOff 'Clear Counters'
      on Press: InvertBit("HmiDb_ClearCounter")
      on Release: InvertBit("HmiDb_ClearCounter")
   Rectangle "Rectangle_8" at 461,318 size 24x22
      Appearance <- "AlreadyFilledSlotArray_Row1Y{0}"
   Rectangle "Rectangle_9" at 431,318 size 24x22
      Appearance <- "AlreadyFilledSlotArray_Row2Y{0}"
   Rectangle "Rectangle_10" at 401,318 size 24x22
      Appearance <- "AlreadyFilledSlotArray_Row3Y{0}"
   Rectangle "Rectangle_11" at 371,318 size 24x22
      Appearance <- "AlreadyFilledSlotArray_Row4Y{0}"
   Rectangle "Rectangle_12" at 341,318 size 24x22
      Appearance <- "AlreadyFilledSlotArray_Row5Y{0}"
   Rectangle "Rectangle_13" at 311,318 size 24x22
      Appearance <- "AlreadyFilledSlotArray_Row6Y{0}"
   Rectangle "Rectangle_14" at 281,318 size 24x22
      Appearance <- "AlreadyFilledSlotArray_Row7Y{0}"
   Rectangle "Rectangle_15" at 251,318 size 24x22
      Appearance <- "AlreadyFilledSlotArray_Row8Y{0}"
   Rectangle "Rectangle_16" at 222,318 size 24x22
      Appearance <- "AlreadyFilledSlotArray_Row9Y{0}"
   Rectangle "Rectangle_17" at 461,286 size 24x22
      Appearance <- "AlreadyFilledSlotArray_Row1Y{1}"
   Rectangle "Rectangle_18" at 431,286 size 24x22
      Appearance <- "AlreadyFilledSlotArray_Row2Y{1}"
   Rectangle "Rectangle_19" at 401,286 size 24x22
      Appearance <- "AlreadyFilledSlotArray_Row3Y{1}"
   Rectangle "Rectangle_20" at 371,286 size 24x22
      Appearance <- "AlreadyFilledSlotArray_Row4Y{1}"
   Rectangle "Rectangle_21" at 341,286 size 24x22
      Appearance <- "AlreadyFilledSlotArray_Row5Y{1}"
   Rectangle "Rectangle_22" at 311,286 size 24x22
      Appearance <- "AlreadyFilledSlotArray_Row6Y{1}"
   Rectangle "Rectangle_23" at 281,286 size 24x22
      Appearance <- "AlreadyFilledSlotArray_Row7Y{1}"
   Rectangle "Rectangle_24" at 251,286 size 24x22
      Appearance <- "AlreadyFilledSlotArray_Row8Y{1}"
   Rectangle "Rectangle_25" at 222,286 size 24x22
      Appearance <- "AlreadyFilledSlotArray_Row9Y{1}"
   Rectangle "Rectangle_26" at 461,253 size 24x22
      Appearance <- "AlreadyFilledSlotArray_Row1Y{2}"
   Rectangle "Rectangle_27" at 431,253 size 24x22
      Appearance <- "AlreadyFilledSlotArray_Row2Y{2}"
   Rectangle "Rectangle_28" at 401,253 size 24x22
      Appearance <- "AlreadyFilledSlotArray_Row3Y{2}"
   Rectangle "Rectangle_29" at 371,253 size 24x22
      Appearance <- "AlreadyFilledSlotArray_Row4Y{2}"
   Rectangle "Rectangle_30" at 341,253 size 24x22
      Appearance <- "AlreadyFilledSlotArray_Row5Y{2}"
   Rectangle "Rectangle_31" at 311,253 size 24x22
      Appearance <- "AlreadyFilledSlotArray_Row6Y{2}"
   Rectangle "Rectangle_32" at 281,253 size 24x22
      Appearance <- "AlreadyFilledSlotArray_Row7Y{2}"
   Rectangle "Rectangle_33" at 251,253 size 24x22
      Appearance <- "AlreadyFilledSlotArray_Row8Y{2}"
   Rectangle "Rectangle_34" at 222,253 size 24x22
      Appearance <- "AlreadyFilledSlotArray_Row9Y{2}"
   Rectangle "Rectangle_35" at 461,220 size 24x22
      Appearance <- "AlreadyFilledSlotArray_Row1Y{3}"
   Rectangle "Rectangle_36" at 431,220 size 24x22
      Appearance <- "AlreadyFilledSlotArray_Row2Y{3}"
   Rectangle "Rectangle_37" at 401,220 size 24x22
      Appearance <- "AlreadyFilledSlotArray_Row3Y{3}"
   Rectangle "Rectangle_38" at 371,220 size 24x22
      Appearance <- "AlreadyFilledSlotArray_Row4Y{3}"
   Rectangle "Rectangle_39" at 341,220 size 24x22
      Appearance <- "AlreadyFilledSlotArray_Row5Y{3}"
   Rectangle "Rectangle_40" at 311,220 size 24x22
      Appearance <- "AlreadyFilledSlotArray_Row6Y{3}"
   Rectangle "Rectangle_41" at 281,220 size 24x22
      Appearance <- "AlreadyFilledSlotArray_Row7Y{3}"
   Rectangle "Rectangle_42" at 251,220 size 24x22
      Appearance <- "AlreadyFilledSlotArray_Row8Y{3}"
   Rectangle "Rectangle_43" at 222,220 size 24x22
      Appearance <- "AlreadyFilledSlotArray_Row9Y{3}"
   Rectangle "Rectangle_44" at 461,186 size 24x22
      Appearance <- "AlreadyFilledSlotArray_Row1Y{4}"
   Rectangle "Rectangle_45" at 431,186 size 24x22
      Appearance <- "AlreadyFilledSlotArray_Row2Y{4}"
   Rectangle "Rectangle_46" at 401,186 size 24x22
      Appearance <- "AlreadyFilledSlotArray_Row3Y{4}"
   Rectangle "Rectangle_47" at 371,186 size 24x22
      Appearance <- "AlreadyFilledSlotArray_Row4Y{4}"
   Rectangle "Rectangle_48" at 341,186 size 24x22
      Appearance <- "AlreadyFilledSlotArray_Row5Y{4}"
   Rectangle "Rectangle_49" at 311,186 size 24x22
      Appearance <- "AlreadyFilledSlotArray_Row6Y{4}"
   Rectangle "Rectangle_50" at 281,186 size 24x22
      Appearance <- "AlreadyFilledSlotArray_Row7Y{4}"
   Rectangle "Rectangle_51" at 251,186 size 24x22
      Appearance <- "AlreadyFilledSlotArray_Row8Y{4}"
   Rectangle "Rectangle_52" at 222,186 size 24x22
      Appearance <- "AlreadyFilledSlotArray_Row9Y{4}"
   Rectangle "Rectangle_53" at 461,152 size 24x22
      Appearance <- "AlreadyFilledSlotArray_Row1Y{5}"
   Rectangle "Rectangle_54" at 431,152 size 24x22
      Appearance <- "AlreadyFilledSlotArray_Row2Y{5}"
   Rectangle "Rectangle_55" at 401,152 size 24x22
      Appearance <- "AlreadyFilledSlotArray_Row3Y{5}"
   Rectangle "Rectangle_56" at 371,152 size 24x22
      Appearance <- "AlreadyFilledSlotArray_Row4Y{5}"
   Rectangle "Rectangle_57" at 341,152 size 24x22
      Appearance <- "AlreadyFilledSlotArray_Row5Y{5}"
   Rectangle "Rectangle_58" at 311,152 size 24x22
      Appearance <- "AlreadyFilledSlotArray_Row6Y{5}"
   Rectangle "Rectangle_59" at 281,152 size 24x22
      Appearance <- "AlreadyFilledSlotArray_Row7Y{5}"
   Rectangle "Rectangle_60" at 251,152 size 24x22
      Appearance <- "AlreadyFilledSlotArray_Row8Y{5}"
   Rectangle "Rectangle_61" at 222,152 size 24x22
      Appearance <- "AlreadyFilledSlotArray_Row9Y{5}"

screen "CalibrateCrane" 800x600
   SymbolicIOField "Symbolic I/O field_1" at 595,8 size 170x32; TextOn '1'; TextOff '0'; TextList "scadascreenlist"
      on Change: ActivateScreenByNumber("THEscreen", 2)
      ProcessValue <- "THEscreen"
   SymbolicIOField "Symbolic I/O field_2" at 543,165 size 129x32; TextOff '0'; TextOn '1'; TextList "ZarrayList"
      ProcessValue <- "ylist"
   SymbolicIOField "Symbolic I/O field_3" at 381,166 size 137x32; TextOn '1'; TextOff '0'; TextList "XarrayList"
      ProcessValue <- "xlist"
   TextField "Text field_1" at 590,111 size 21x34; Text 'Z'
   TextField "Text field_2" at 439,113 size 22x34; Text 'X'
   IOField "I/O field_1" at 560,503 size 118x32; FormatPattern 99999
      ProcessValue <- "HmiDb_CalInputVal"
   TextField "Text field_3" at 560,476 size 81x22; Text 'Insert MM'
   Button "Button_1" at 695,503 size 96x32; TextOff 'Save X'
      on Press: InvertBit("HmiDb_HmiSaveArmCal")
      on Release: InvertBit("HmiDb_HmiSaveArmCal")
   Button "Button_2" at 695,546 size 96x32; TextOff 'Save Y'
      on Press: InvertBit("HmiDb_HmiSaveArmCalY")
      on Release: InvertBit("HmiDb_HmiSaveArmCalY")
   IOField "I/O field_2" at 387,503 size 96x32; FormatPattern 9999
      ProcessValue <- "HmiDb_CurrentPositionY"
   IOField "I/O field_3" at 283,503 size 96x32; FormatPattern 99999
      ProcessValue <- "HmiDb_CurrentPositionX"
   TextField "Text field_4" at 288,474 size 40x22; Text 'DB X'
   TextField "Text field_5" at 392,474 size 39x22; Text 'DB Z'
   IOField "I/O field_4" at 387,563 size 96x32; FormatPattern 9999
      ProcessValue <- "OutputsDB_CraneOutput_Ymm"
   IOField "I/O field_5" at 283,563 size 96x32; FormatPattern 99999
      ProcessValue <- "OutputsDB_CraneOutput_Xmm"
   TextField "Text field_6" at 288,534 size 63x22; Text 'Crane X'
   TextField "Text field_7" at 392,534 size 62x22; Text 'Crane Z'
   Slider "Slider_2" at 57,48 size 60x525; Caption 'SIMATIC'
      ProcessValue <- "jogmodeDB_CraneXjog"
   Slider "Slider_1" at 171,49 size 60x526; Caption 'SIMATIC'
      ProcessValue <- "jogmodeDB_CraneYjog"
   TextField "Text field_8" at 73,7 size 22x34; Text 'X'
   TextField "Text field_9" at 186,8 size 21x34; Text 'Z'
   Button "Button_9" at 378,246 size 296x32; TextOff 'Calibrate Mode'
      on Deactivate: SetTag("jogmodeDB_CraneXjog", 0); SetTag("jogmodeDB_CraneYjog", 0)
      on Click: InvertBit("Modes_Modes_JogMode")
      on Activate: SetTag("jogmodeDB_CraneXjog", 0); SetTag("jogmodeDB_CraneYjog", 0)
      Appearance <- "Modes_Modes_JogMode"
   Button "Button_3" at 441,371 size 35x32; TextOff '10'
      on Press: SetTag("InputsDB_AdjustX", 10); SetBit("InputsDB_PressAdjustX")
      on Release: SetTag("InputsDB_AdjustX", 0); ResetBit("InputsDB_PressAdjustX")
   Button "Button_4" at 472,371 size 35x32; TextOff '1'
      on Press: SetTag("InputsDB_AdjustX", 1); SetBit("InputsDB_PressAdjustX")
      on Release: SetTag("InputsDB_AdjustX", 0); ResetBit("InputsDB_PressAdjustX")
   Button "Button_5" at 505,311 size 35x32; TextOff '10'
      on Release: SetTag("InputsDB_AdjustY", 0); ResetBit("InputsDB_PressAdjustY")
      on Press: SetTag("InputsDB_AdjustY", 10); SetBit("InputsDB_PressAdjustY")
   Button "Button_6" at 505,340 size 35x32; TextOff '1'
      on Release: SetTag("InputsDB_AdjustY", 0); ResetBit("InputsDB_PressAdjustY")
      on Press: SetTag("InputsDB_AdjustY", 1); SetBit("InputsDB_PressAdjustY")
   Button "Button_7" at 505,434 size 35x32; TextOff '10'
      on Release: SetTag("InputsDB_AdjustY", 0); ResetBit("InputsDB_PressAdjustY")
      on Press: SetTag("InputsDB_AdjustY", -10); SetBit("InputsDB_PressAdjustY")
   Button "Button_8" at 505,402 size 35x32; TextOff '1'
      on Release: SetTag("InputsDB_AdjustY", 0); ResetBit("InputsDB_PressAdjustY")
      on Press: SetTag("InputsDB_AdjustY", -1); SetBit("InputsDB_PressAdjustY")
   Button "Button_10" at 506,371 size 35x32; TextOff 'Text'
   Button "Button_11" at 573,371 size 35x32; TextOff '10'
      on Release: SetTag("InputsDB_AdjustX", 0); ResetBit("InputsDB_PressAdjustX")
      on Press: SetTag("InputsDB_AdjustX", -10); SetBit("InputsDB_PressAdjustX")
   Button "Button_12" at 540,371 size 35x32; TextOff '1'
      on Release: SetTag("InputsDB_AdjustX", 0); ResetBit("InputsDB_PressAdjustX")
      on Press: SetTag("InputsDB_AdjustX", -1); SetBit("InputsDB_PressAdjustX")

PopupScreen "Pop-up screen_1" 240x240
   TextField "Text field_1" at 71,52 size 80x22; Text 'You sure?'
   Button "Button_1" at 11,127 size 96x32; TextOff 'yes'
      on Press: function_efd93a16("Pop-up screen_1", 0, 0, -1, -1, 1); InvertBit("HmiDb_ClearStock")
      on Release: InvertBit("HmiDb_ClearStock")
   Button "Button_2" at 124,129 size 96x32; TextOff 'no'
      on Press: function_efd93a16("Pop-up screen_1", 0, 0, -1, -1, 1)
*)